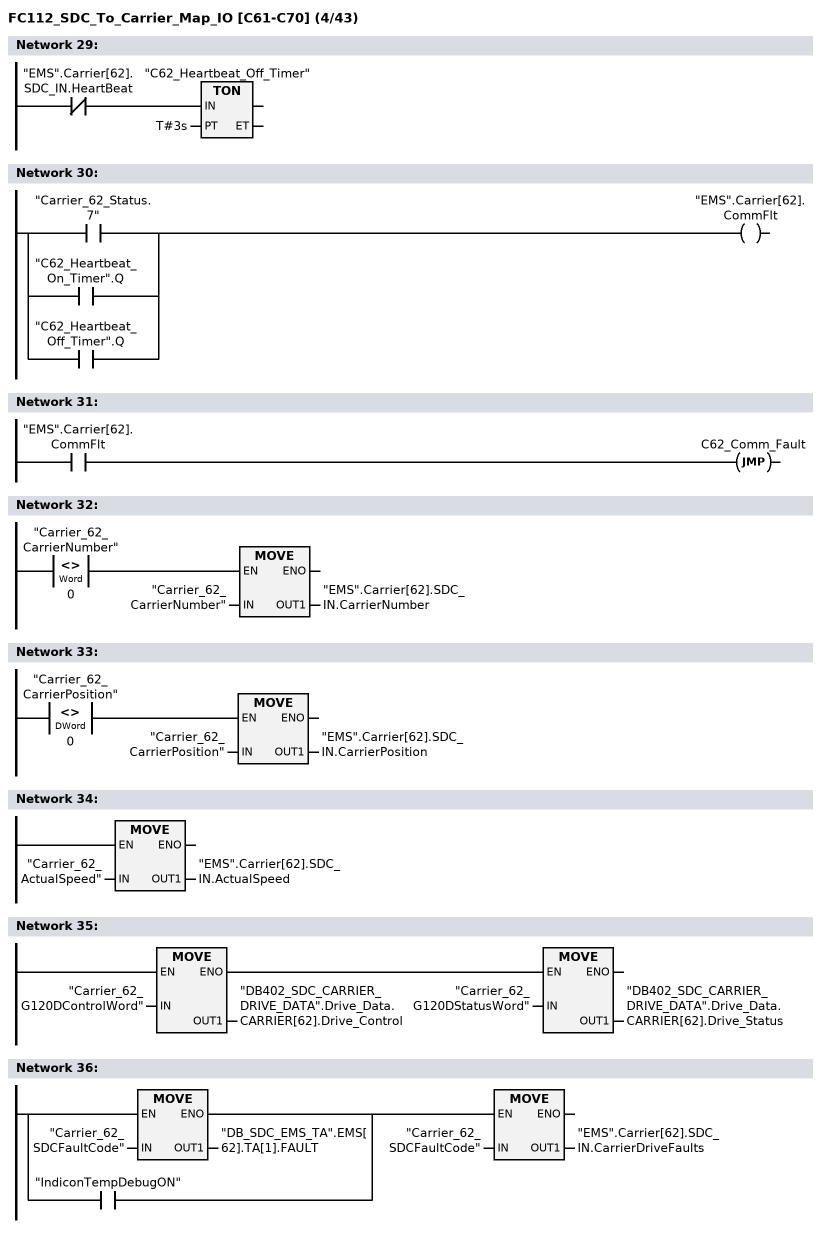
   "C62_Heartbeat_Off_Timer".TON(IN := NOT "EMS".Carrier[62].SDC_IN.HeartBeat, PT := T#3s);
END_REGION

REGION Network 30
   RUNG wire#powerrail
      Contact( "Carrier_62_Status.7" )
      wire#w1
      Coil( "EMS".Carrier[62].CommFlt )
   END_RUNG
   RUNG wire#powerrail
      Contact( "C62_Heartbeat_On_Timer".Q )
   END_RUNG wire#w1
   RUNG wire#powerrail
      Contact( "C62_Heartbeat_Off_Timer".Q )
   END_RUNG wire#w1
   // the same network as SCL:
   "EMS".Carrier[62].CommFlt := "Carrier_62_Status.7" OR "C62_Heartbeat_On_Timer".Q OR "C62_Heartbeat_Off_Timer".Q;
END_REGION

REGION Network 31
   RUNG wire#powerrail
      Contact( "EMS".Carrier[62].CommFlt )
      JumpCoil( C62_Comm_Fault )
   END_RUNG
   // the same network as SCL:
   IF "EMS".Carrier[62].CommFlt THEN GOTO C62_Comm_Fault; END_IF;
END_REGION

REGION Network 32
   RUNG wire#powerrail
      { S7_Templates := "SrcType := Word" } NE_Contact(in1 := "Carrier_62_CarrierNumber", in2 := 0)
      Move(in := "Carrier_62_CarrierNumber", out1 => "EMS".Carrier[62].SDC_IN.CarrierNumber)
   END_RUNG
   // the same network as SCL:
   IF "Carrier_62_CarrierNumber" <> 0 THEN
       "EMS".Carrier[62].SDC_IN.CarrierNumber := "Carrier_62_CarrierNumber";
   END_IF;
END_REGION

REGION Network 33
   RUNG wire#powerrail
      { S7_Templates := "SrcType := DWord" } NE_Contact(in1 := "Carrier_62_CarrierPosition", in2 := 0)
      Move(in := "Carrier_62_CarrierPosition", out1 => "EMS".Carrier[62].SDC_IN.CarrierPosition)
   END_RUNG
   // the same network as SCL:
   IF "Carrier_62_CarrierPosition" <> 0 THEN
       "EMS".Carrier[62].SDC_IN.CarrierPosition := "Carrier_62_CarrierPosition";
   END_IF;
END_REGION

REGION Network 34
   RUNG wire#powerrail
      Move(in := "Carrier_62_ActualSpeed", out1 => "EMS".Carrier[62].SDC_IN.ActualSpeed)
   END_RUNG
   // the same network as SCL:
   "EMS".Carrier[62].SDC_IN.ActualSpeed := "Carrier_62_ActualSpeed";
END_REGION

REGION Network 35
   RUNG wire#powerrail
      Move(in := "Carrier_62_G120DControlWord", out1 => "DB402_SDC_CARRIER_DRIVE_DATA".Drive_Data.CARRIER[62].Drive_Control)
      Move(in := "Carrier_62_G120DStatusWord", out1 => "DB402_SDC_CARRIER_DRIVE_DATA".Drive_Data.CARRIER[62].Drive_Status)
   END_RUNG
   // the same network as SCL:
   "DB402_SDC_CARRIER_DRIVE_DATA".Drive_Data.CARRIER[62].Drive_Control := "Carrier_62_G120DControlWord";
   "DB402_SDC_CARRIER_DRIVE_DATA".Drive_Data.CARRIER[62].Drive_Status := "Carrier_62_G120DStatusWord";
END_REGION

REGION Network 36
   RUNG wire#powerrail
      Move(in := "Carrier_62_SDCFaultCode", out1 => "DB_SDC_EMS_TA".EMS[62].TA[1].FAULT)
      wire#w1
      Move(in := "Carrier_62_SDCFaultCode", out1 => "EMS".Carrier[62].SDC_IN.CarrierDriveFaults)
   END_RUNG
   RUNG wire#powerrail
      Contact( "IndiconTempDebugON" )
   END_RUNG wire#w1
   // the same network as SCL:
   "DB_SDC_EMS_TA".EMS[62].TA[1].FAULT := "Carrier_62_SDCFaultCode";
   IF TRUE OR "IndiconTempDebugON" THEN
       "EMS".Carrier[62].SDC_IN.CarrierDriveFaults := "Carrier_62_SDCFaultCode";
   END_IF;
END_REGION

REGION Network 37
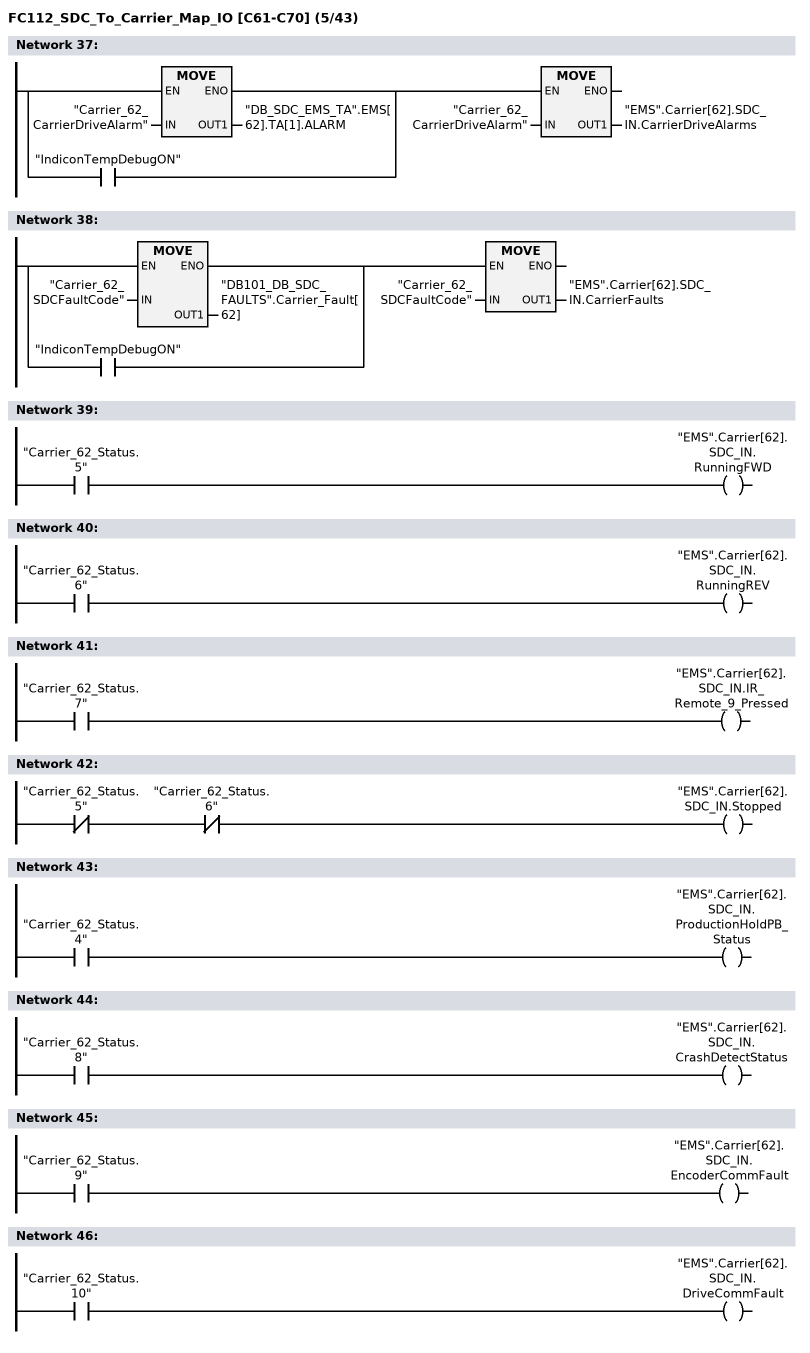
   RUNG wire#powerrail
      Move(in := "Carrier_62_CarrierDriveAlarm", out1 => "DB_SDC_EMS_TA".EMS[62].TA[1].ALARM)
      wire#w1
      Move(in := "Carrier_62_CarrierDriveAlarm", out1 => "EMS".Carrier[62].SDC_IN.CarrierDriveAlarms)
   END_RUNG
   RUNG wire#powerrail
      Contact( "IndiconTempDebugON" )
   END_RUNG wire#w1
   // the same network as SCL:
   "DB_SDC_EMS_TA".EMS[62].TA[1].ALARM := "Carrier_62_CarrierDriveAlarm";
   IF TRUE OR "IndiconTempDebugON" THEN
       "EMS".Carrier[62].SDC_IN.CarrierDriveAlarms := "Carrier_62_CarrierDriveAlarm";
   END_IF;
END_REGION

REGION Network 38
   RUNG wire#powerrail
      Move(in := "Carrier_62_SDCFaultCode", out1 => "DB101_DB_SDC_FAULTS".Carrier_Fault[62])
      wire#w1
      Move(in := "Carrier_62_SDCFaultCode", out1 => "EMS".Carrier[62].SDC_IN.CarrierFaults)
   END_RUNG
   RUNG wire#powerrail
      Contact( "IndiconTempDebugON" )
   END_RUNG wire#w1
   // the same network as SCL:
   "DB101_DB_SDC_FAULTS".Carrier_Fault[62] := "Carrier_62_SDCFaultCode";
   IF TRUE OR "IndiconTempDebugON" THEN
       "EMS".Carrier[62].SDC_IN.CarrierFaults := "Carrier_62_SDCFaultCode";
   END_IF;
END_REGION

REGION Network 39
   RUNG wire#powerrail
      Contact( "Carrier_62_Status.5" )
      Coil( "EMS".Carrier[62].SDC_IN.RunningFWD )
   END_RUNG
   // the same network as SCL:
   "EMS".Carrier[62].SDC_IN.RunningFWD := "Carrier_62_Status.5";
END_REGION

REGION Network 40
   RUNG wire#powerrail
      Contact( "Carrier_62_Status.6" )
      Coil( "EMS".Carrier[62].SDC_IN.RunningREV )
   END_RUNG
   // the same network as SCL:
   "EMS".Carrier[62].SDC_IN.RunningREV := "Carrier_62_Status.6";
END_REGION

REGION Network 41
   RUNG wire#powerrail
      Contact( "Carrier_62_Status.7" )
      Coil( "EMS".Carrier[62].SDC_IN.IR_Remote_9_Pressed )
   END_RUNG
   // the same network as SCL:
   "EMS".Carrier[62].SDC_IN.IR_Remote_9_Pressed := "Carrier_62_Status.7";
END_REGION

REGION Network 42
   RUNG wire#powerrail
      I_Contact( "Carrier_62_Status.5" )
      I_Contact( "Carrier_62_Status.6" )
      Coil( "EMS".Carrier[62].SDC_IN.Stopped )
   END_RUNG
   // the same network as SCL:
   "EMS".Carrier[62].SDC_IN.Stopped := NOT "Carrier_62_Status.5" AND NOT "Carrier_62_Status.6";
END_REGION

REGION Network 43
   RUNG wire#powerrail
      Contact( "Carrier_62_Status.4" )
      Coil( "EMS".Carrier[62].SDC_IN.ProductionHoldPB_Status )
   END_RUNG
   // the same network as SCL:
   "EMS".Carrier[62].SDC_IN.ProductionHoldPB_Status := "Carrier_62_Status.4";
END_REGION

REGION Network 44
   RUNG wire#powerrail
      Contact( "Carrier_62_Status.8" )
      Coil( "EMS".Carrier[62].SDC_IN.CrashDetectStatus )
   END_RUNG
   // the same network as SCL:
   "EMS".Carrier[62].SDC_IN.CrashDetectStatus := "Carrier_62_Status.8";
END_REGION

REGION Network 45
   RUNG wire#powerrail
      Contact( "Carrier_62_Status.9" )
      Coil( "EMS".Carrier[62].SDC_IN.EncoderCommFault )
   END_RUNG
   // the same network as SCL:
   "EMS".Carrier[62].SDC_IN.EncoderCommFault := "Carrier_62_Status.9";
END_REGION

REGION Network 46
   RUNG wire#powerrail
      Contact( "Carrier_62_Status.10" )
      Coil( "EMS".Carrier[62].SDC_IN.DriveCommFault )
   END_RUNG
   // the same network as SCL:
   "EMS".Carrier[62].SDC_IN.DriveCommFault := "Carrier_62_Status.10";
END_REGION

REGION Network 47
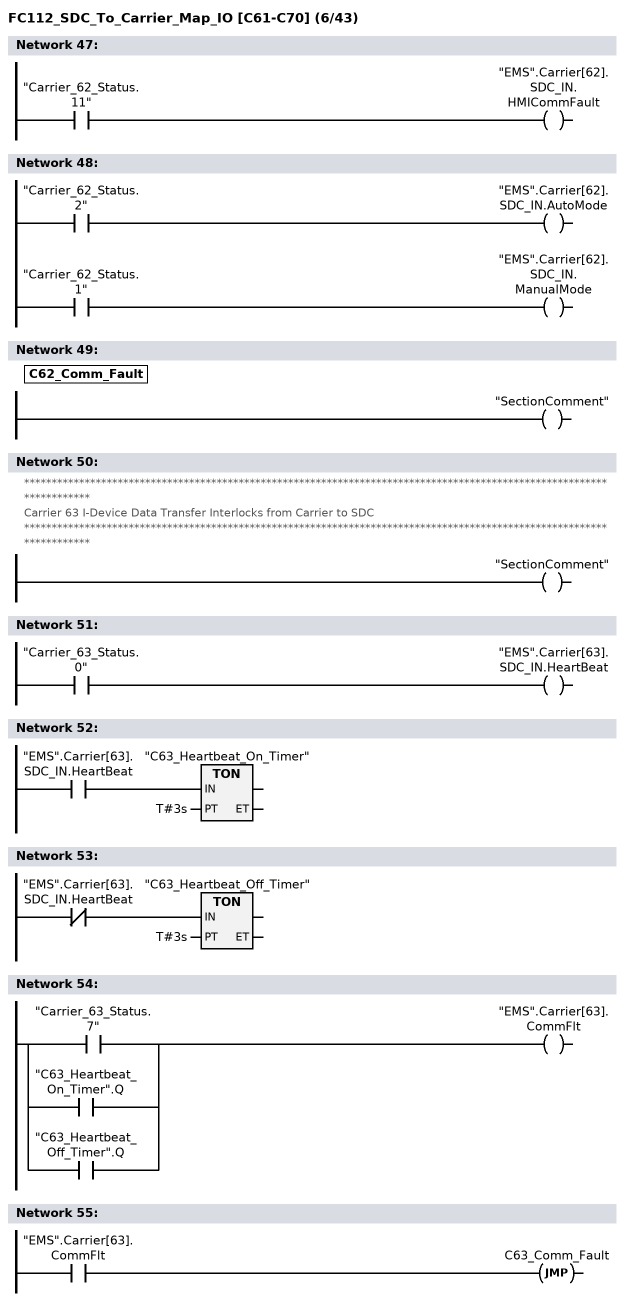
   RUNG wire#powerrail
      Contact( "Carrier_62_Status.11" )
      Coil( "EMS".Carrier[62].SDC_IN.HMICommFault )
   END_RUNG
   // the same network as SCL:
   "EMS".Carrier[62].SDC_IN.HMICommFault := "Carrier_62_Status.11";
END_REGION

REGION Network 48
   RUNG wire#powerrail
      Contact( "Carrier_62_Status.2" )
      Coil( "EMS".Carrier[62].SDC_IN.AutoMode )
   END_RUNG
   RUNG wire#powerrail
      Contact( "Carrier_62_Status.1" )
      Coil( "EMS".Carrier[62].SDC_IN.ManualMode )
   END_RUNG
   // the same network as SCL:
   "EMS".Carrier[62].SDC_IN.AutoMode := "Carrier_62_Status.2";
   "EMS".Carrier[62].SDC_IN.ManualMode := "Carrier_62_Status.1";
END_REGION

REGION Network 49
   Label( C62_Comm_Fault )
   RUNG wire#powerrail
      Coil( "SectionComment" )
   END_RUNG
   // the same network as SCL:
   C62_Comm_Fault:
   "SectionComment" := TRUE;
END_REGION

REGION Network 50
   // **********************************************************************************************************************
   // 
   // Carrier 63 I-Device Data Transfer Interlocks from Carrier to SDC
   // 
   // **********************************************************************************************************************
   RUNG wire#powerrail
      Coil( "SectionComment" )
   END_RUNG
   // the same network as SCL:
   "SectionComment" := TRUE;
END_REGION

REGION Network 51
   RUNG wire#powerrail
      Contact( "Carrier_63_Status.0" )
      Coil( "EMS".Carrier[63].SDC_IN.HeartBeat )
   END_RUNG
   // the same network as SCL:
   "EMS".Carrier[63].SDC_IN.HeartBeat := "Carrier_63_Status.0";
END_REGION

REGION Network 52
   "C63_Heartbeat_On_Timer".TON(IN := "EMS".Carrier[63].SDC_IN.HeartBeat, PT := T#3s);
END_REGION

REGION Network 53
   "C63_Heartbeat_Off_Timer".TON(IN := NOT "EMS".Carrier[63].SDC_IN.HeartBeat, PT := T#3s);
END_REGION

REGION Network 54
   RUNG wire#powerrail
      Contact( "Carrier_63_Status.7" )
      wire#w1
      Coil( "EMS".Carrier[63].CommFlt )
   END_RUNG
   RUNG wire#powerrail
      Contact( "C63_Heartbeat_On_Timer".Q )
   END_RUNG wire#w1
   RUNG wire#powerrail
      Contact( "C63_Heartbeat_Off_Timer".Q )
   END_RUNG wire#w1
   // the same network as SCL:
   "EMS".Carrier[63].CommFlt := "Carrier_63_Status.7" OR "C63_Heartbeat_On_Timer".Q OR "C63_Heartbeat_Off_Timer".Q;
END_REGION

REGION Network 55
   RUNG wire#powerrail
      Contact( "EMS".Carrier[63].CommFlt )
      JumpCoil( C63_Comm_Fault )
   END_RUNG
   // the same network as SCL:
   IF "EMS".Carrier[63].CommFlt THEN GOTO C63_Comm_Fault; END_IF;
END_REGION

REGION Network 56
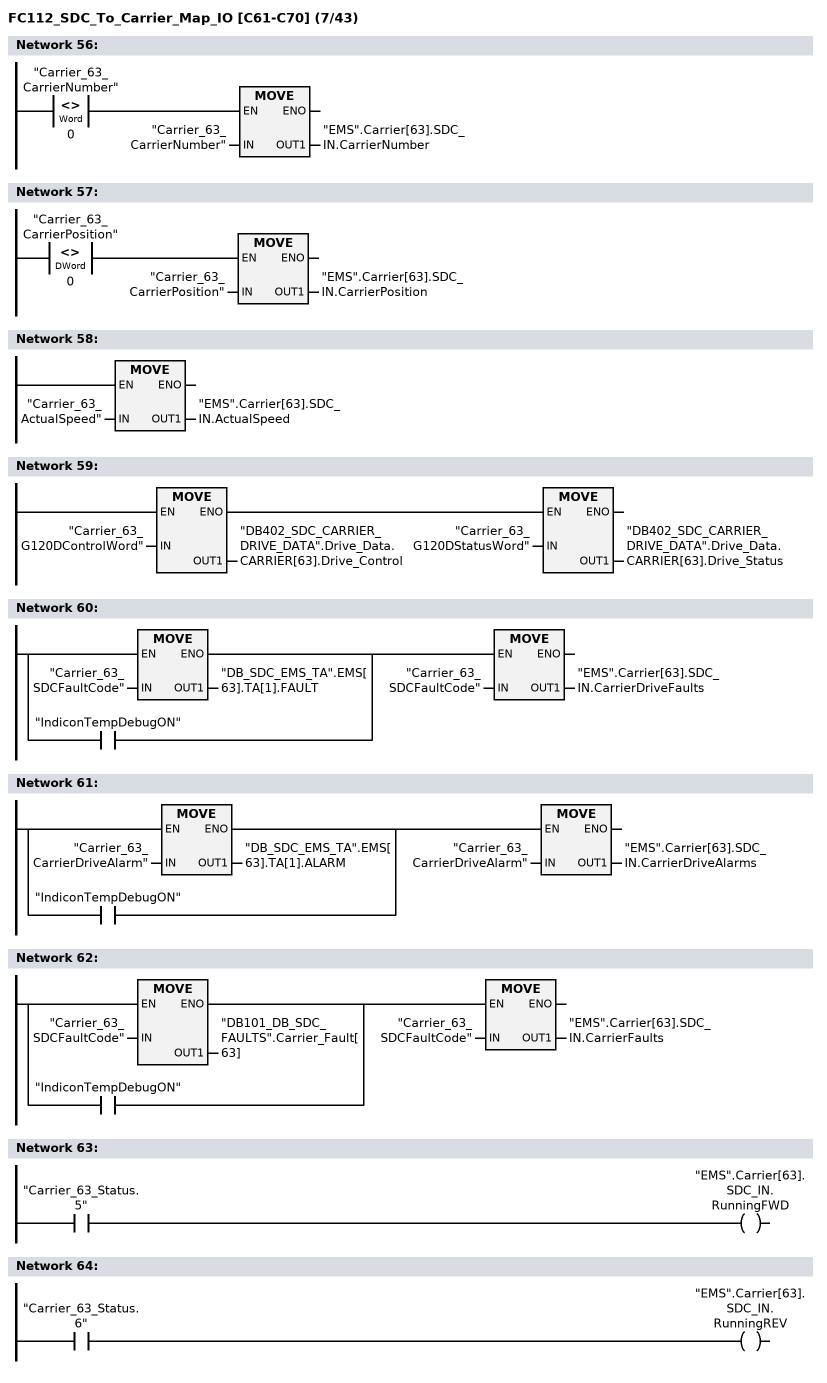
   RUNG wire#powerrail
      { S7_Templates := "SrcType := Word" } NE_Contact(in1 := "Carrier_63_CarrierNumber", in2 := 0)
      Move(in := "Carrier_63_CarrierNumber", out1 => "EMS".Carrier[63].SDC_IN.CarrierNumber)
   END_RUNG
   // the same network as SCL:
   IF "Carrier_63_CarrierNumber" <> 0 THEN
       "EMS".Carrier[63].SDC_IN.CarrierNumber := "Carrier_63_CarrierNumber";
   END_IF;
END_REGION

REGION Network 57
   RUNG wire#powerrail
      { S7_Templates := "SrcType := DWord" } NE_Contact(in1 := "Carrier_63_CarrierPosition", in2 := 0)
      Move(in := "Carrier_63_CarrierPosition", out1 => "EMS".Carrier[63].SDC_IN.CarrierPosition)
   END_RUNG
   // the same network as SCL:
   IF "Carrier_63_CarrierPosition" <> 0 THEN
       "EMS".Carrier[63].SDC_IN.CarrierPosition := "Carrier_63_CarrierPosition";
   END_IF;
END_REGION

REGION Network 58
   RUNG wire#powerrail
      Move(in := "Carrier_63_ActualSpeed", out1 => "EMS".Carrier[63].SDC_IN.ActualSpeed)
   END_RUNG
   // the same network as SCL:
   "EMS".Carrier[63].SDC_IN.ActualSpeed := "Carrier_63_ActualSpeed";
END_REGION

REGION Network 59
   RUNG wire#powerrail
      Move(in := "Carrier_63_G120DControlWord", out1 => "DB402_SDC_CARRIER_DRIVE_DATA".Drive_Data.CARRIER[63].Drive_Control)
      Move(in := "Carrier_63_G120DStatusWord", out1 => "DB402_SDC_CARRIER_DRIVE_DATA".Drive_Data.CARRIER[63].Drive_Status)
   END_RUNG
   // the same network as SCL:
   "DB402_SDC_CARRIER_DRIVE_DATA".Drive_Data.CARRIER[63].Drive_Control := "Carrier_63_G120DControlWord";
   "DB402_SDC_CARRIER_DRIVE_DATA".Drive_Data.CARRIER[63].Drive_Status := "Carrier_63_G120DStatusWord";
END_REGION

REGION Network 60
   RUNG wire#powerrail
      Move(in := "Carrier_63_SDCFaultCode", out1 => "DB_SDC_EMS_TA".EMS[63].TA[1].FAULT)
      wire#w1
      Move(in := "Carrier_63_SDCFaultCode", out1 => "EMS".Carrier[63].SDC_IN.CarrierDriveFaults)
   END_RUNG
   RUNG wire#powerrail
      Contact( "IndiconTempDebugON" )
   END_RUNG wire#w1
   // the same network as SCL:
   "DB_SDC_EMS_TA".EMS[63].TA[1].FAULT := "Carrier_63_SDCFaultCode";
   IF TRUE OR "IndiconTempDebugON" THEN
       "EMS".Carrier[63].SDC_IN.CarrierDriveFaults := "Carrier_63_SDCFaultCode";
   END_IF;
END_REGION

REGION Network 61
   RUNG wire#powerrail
      Move(in := "Carrier_63_CarrierDriveAlarm", out1 => "DB_SDC_EMS_TA".EMS[63].TA[1].ALARM)
      wire#w1
      Move(in := "Carrier_63_CarrierDriveAlarm", out1 => "EMS".Carrier[63].SDC_IN.CarrierDriveAlarms)
   END_RUNG
   RUNG wire#powerrail
      Contact( "IndiconTempDebugON" )
   END_RUNG wire#w1
   // the same network as SCL:
   "DB_SDC_EMS_TA".EMS[63].TA[1].ALARM := "Carrier_63_CarrierDriveAlarm";
   IF TRUE OR "IndiconTempDebugON" THEN
       "EMS".Carrier[63].SDC_IN.CarrierDriveAlarms := "Carrier_63_CarrierDriveAlarm";
   END_IF;
END_REGION

REGION Network 62
   RUNG wire#powerrail
      Move(in := "Carrier_63_SDCFaultCode", out1 => "DB101_DB_SDC_FAULTS".Carrier_Fault[63])
      wire#w1
      Move(in := "Carrier_63_SDCFaultCode", out1 => "EMS".Carrier[63].SDC_IN.CarrierFaults)
   END_RUNG
   RUNG wire#powerrail
      Contact( "IndiconTempDebugON" )
   END_RUNG wire#w1
   // the same network as SCL:
   "DB101_DB_SDC_FAULTS".Carrier_Fault[63] := "Carrier_63_SDCFaultCode";
   IF TRUE OR "IndiconTempDebugON" THEN
       "EMS".Carrier[63].SDC_IN.CarrierFaults := "Carrier_63_SDCFaultCode";
   END_IF;
END_REGION

REGION Network 63
   RUNG wire#powerrail
      Contact( "Carrier_63_Status.5" )
      Coil( "EMS".Carrier[63].SDC_IN.RunningFWD )
   END_RUNG
   // the same network as SCL:
   "EMS".Carrier[63].SDC_IN.RunningFWD := "Carrier_63_Status.5";
END_REGION

REGION Network 64
   RUNG wire#powerrail
      Contact( "Carrier_63_Status.6" )
      Coil( "EMS".Carrier[63].SDC_IN.RunningREV )
   END_RUNG
   // the same network as SCL:
   "EMS".Carrier[63].SDC_IN.RunningREV := "Carrier_63_Status.6";
END_REGION

REGION Network 65
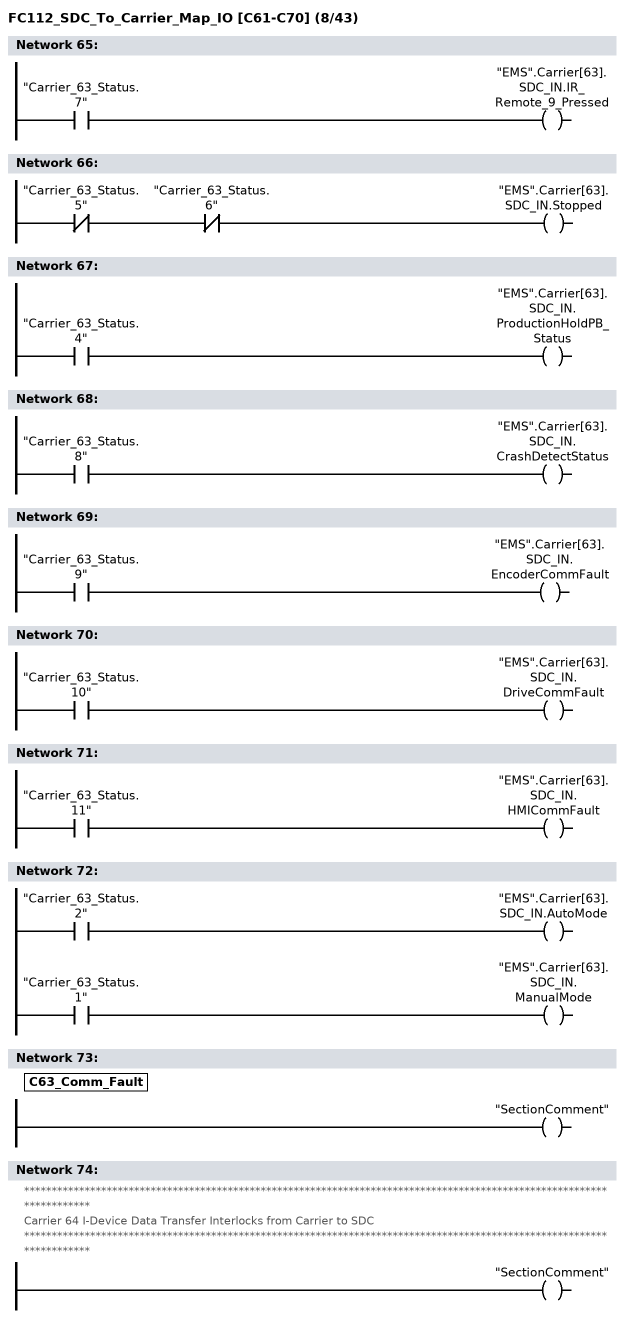
   RUNG wire#powerrail
      Contact( "Carrier_63_Status.7" )
      Coil( "EMS".Carrier[63].SDC_IN.IR_Remote_9_Pressed )
   END_RUNG
   // the same network as SCL:
   "EMS".Carrier[63].SDC_IN.IR_Remote_9_Pressed := "Carrier_63_Status.7";
END_REGION

REGION Network 66
   RUNG wire#powerrail
      I_Contact( "Carrier_63_Status.5" )
      I_Contact( "Carrier_63_Status.6" )
      Coil( "EMS".Carrier[63].SDC_IN.Stopped )
   END_RUNG
   // the same network as SCL:
   "EMS".Carrier[63].SDC_IN.Stopped := NOT "Carrier_63_Status.5" AND NOT "Carrier_63_Status.6";
END_REGION

REGION Network 67
   RUNG wire#powerrail
      Contact( "Carrier_63_Status.4" )
      Coil( "EMS".Carrier[63].SDC_IN.ProductionHoldPB_Status )
   END_RUNG
   // the same network as SCL:
   "EMS".Carrier[63].SDC_IN.ProductionHoldPB_Status := "Carrier_63_Status.4";
END_REGION

REGION Network 68
   RUNG wire#powerrail
      Contact( "Carrier_63_Status.8" )
      Coil( "EMS".Carrier[63].SDC_IN.CrashDetectStatus )
   END_RUNG
   // the same network as SCL:
   "EMS".Carrier[63].SDC_IN.CrashDetectStatus := "Carrier_63_Status.8";
END_REGION

REGION Network 69
   RUNG wire#powerrail
      Contact( "Carrier_63_Status.9" )
      Coil( "EMS".Carrier[63].SDC_IN.EncoderCommFault )
   END_RUNG
   // the same network as SCL:
   "EMS".Carrier[63].SDC_IN.EncoderCommFault := "Carrier_63_Status.9";
END_REGION

REGION Network 70
   RUNG wire#powerrail
      Contact( "Carrier_63_Status.10" )
      Coil( "EMS".Carrier[63].SDC_IN.DriveCommFault )
   END_RUNG
   // the same network as SCL:
   "EMS".Carrier[63].SDC_IN.DriveCommFault := "Carrier_63_Status.10";
END_REGION

REGION Network 71
   RUNG wire#powerrail
      Contact( "Carrier_63_Status.11" )
      Coil( "EMS".Carrier[63].SDC_IN.HMICommFault )
   END_RUNG
   // the same network as SCL:
   "EMS".Carrier[63].SDC_IN.HMICommFault := "Carrier_63_Status.11";
END_REGION

REGION Network 72
   RUNG wire#powerrail
      Contact( "Carrier_63_Status.2" )
      Coil( "EMS".Carrier[63].SDC_IN.AutoMode )
   END_RUNG
   RUNG wire#powerrail
      Contact( "Carrier_63_Status.1" )
      Coil( "EMS".Carrier[63].SDC_IN.ManualMode )
   END_RUNG
   // the same network as SCL:
   "EMS".Carrier[63].SDC_IN.AutoMode := "Carrier_63_Status.2";
   "EMS".Carrier[63].SDC_IN.ManualMode := "Carrier_63_Status.1";
END_REGION

REGION Network 73
   Label( C63_Comm_Fault )
   RUNG wire#powerrail
      Coil( "SectionComment" )
   END_RUNG
   // the same network as SCL:
   C63_Comm_Fault:
   "SectionComment" := TRUE;
END_REGION

REGION Network 74
   // **********************************************************************************************************************
   // 
   // Carrier 64 I-Device Data Transfer Interlocks from Carrier to SDC
   // 
   // **********************************************************************************************************************
   RUNG wire#powerrail
      Coil( "SectionComment" )
   END_RUNG
   // the same network as SCL:
   "SectionComment" := TRUE;
END_REGION

REGION Network 75
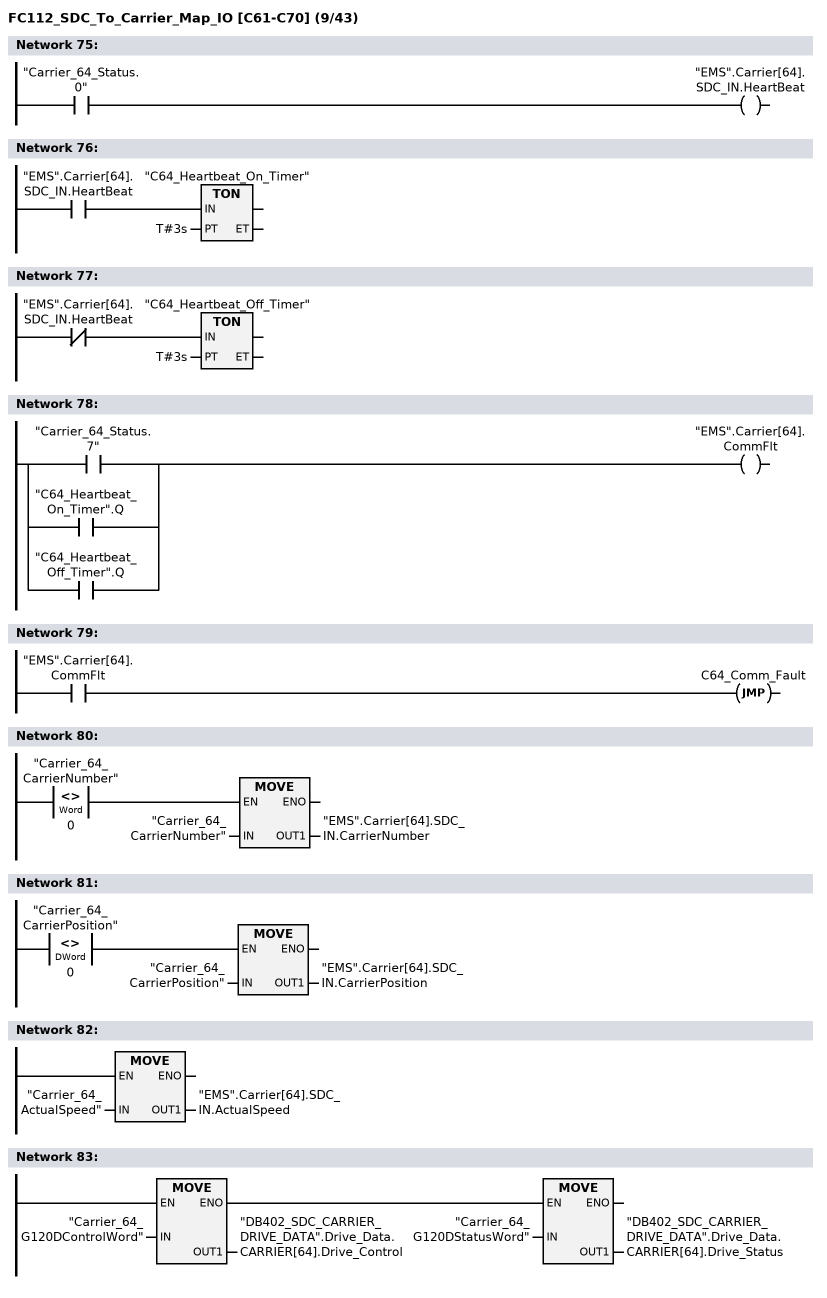
   RUNG wire#powerrail
      Contact( "Carrier_64_Status.0" )
      Coil( "EMS".Carrier[64].SDC_IN.HeartBeat )
   END_RUNG
   // the same network as SCL:
   "EMS".Carrier[64].SDC_IN.HeartBeat := "Carrier_64_Status.0";
END_REGION

REGION Network 76
   "C64_Heartbeat_On_Timer".TON(IN := "EMS".Carrier[64].SDC_IN.HeartBeat, PT := T#3s);
END_REGION

REGION Network 77
   "C64_Heartbeat_Off_Timer".TON(IN := NOT "EMS".Carrier[64].SDC_IN.HeartBeat, PT := T#3s);
END_REGION

REGION Network 78
   RUNG wire#powerrail
      Contact( "Carrier_64_Status.7" )
      wire#w1
      Coil( "EMS".Carrier[64].CommFlt )
   END_RUNG
   RUNG wire#powerrail
      Contact( "C64_Heartbeat_On_Timer".Q )
   END_RUNG wire#w1
   RUNG wire#powerrail
      Contact( "C64_Heartbeat_Off_Timer".Q )
   END_RUNG wire#w1
   // the same network as SCL:
   "EMS".Carrier[64].CommFlt := "Carrier_64_Status.7" OR "C64_Heartbeat_On_Timer".Q OR "C64_Heartbeat_Off_Timer".Q;
END_REGION

REGION Network 79
   RUNG wire#powerrail
      Contact( "EMS".Carrier[64].CommFlt )
      JumpCoil( C64_Comm_Fault )
   END_RUNG
   // the same network as SCL:
   IF "EMS".Carrier[64].CommFlt THEN GOTO C64_Comm_Fault; END_IF;
END_REGION

REGION Network 80
   RUNG wire#powerrail
      { S7_Templates := "SrcType := Word" } NE_Contact(in1 := "Carrier_64_CarrierNumber", in2 := 0)
      Move(in := "Carrier_64_CarrierNumber", out1 => "EMS".Carrier[64].SDC_IN.CarrierNumber)
   END_RUNG
   // the same network as SCL:
   IF "Carrier_64_CarrierNumber" <> 0 THEN
       "EMS".Carrier[64].SDC_IN.CarrierNumber := "Carrier_64_CarrierNumber";
   END_IF;
END_REGION

REGION Network 81
   RUNG wire#powerrail
      { S7_Templates := "SrcType := DWord" } NE_Contact(in1 := "Carrier_64_CarrierPosition", in2 := 0)
      Move(in := "Carrier_64_CarrierPosition", out1 => "EMS".Carrier[64].SDC_IN.CarrierPosition)
   END_RUNG
   // the same network as SCL:
   IF "Carrier_64_CarrierPosition" <> 0 THEN
       "EMS".Carrier[64].SDC_IN.CarrierPosition := "Carrier_64_CarrierPosition";
   END_IF;
END_REGION

REGION Network 82
   RUNG wire#powerrail
      Move(in := "Carrier_64_ActualSpeed", out1 => "EMS".Carrier[64].SDC_IN.ActualSpeed)
   END_RUNG
   // the same network as SCL:
   "EMS".Carrier[64].SDC_IN.ActualSpeed := "Carrier_64_ActualSpeed";
END_REGION

REGION Network 83
   RUNG wire#powerrail
      Move(in := "Carrier_64_G120DControlWord", out1 => "DB402_SDC_CARRIER_DRIVE_DATA".Drive_Data.CARRIER[64].Drive_Control)
      Move(in := "Carrier_64_G120DStatusWord", out1 => "DB402_SDC_CARRIER_DRIVE_DATA".Drive_Data.CARRIER[64].Drive_Status)
   END_RUNG
   // the same network as SCL:
   "DB402_SDC_CARRIER_DRIVE_DATA".Drive_Data.CARRIER[64].Drive_Control := "Carrier_64_G120DControlWord";
   "DB402_SDC_CARRIER_DRIVE_DATA".Drive_Data.CARRIER[64].Drive_Status := "Carrier_64_G120DStatusWord";
END_REGION

REGION Network 84
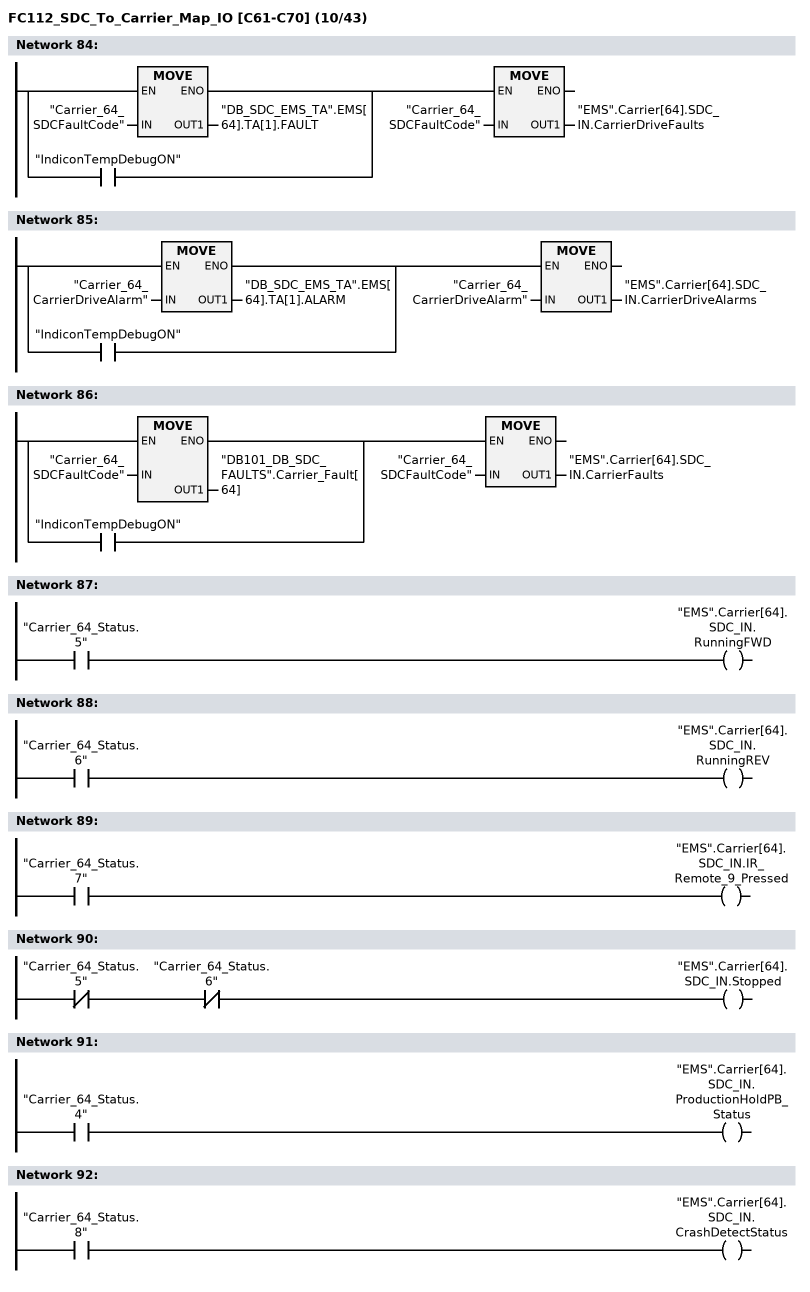
   RUNG wire#powerrail
      Move(in := "Carrier_64_SDCFaultCode", out1 => "DB_SDC_EMS_TA".EMS[64].TA[1].FAULT)
      wire#w1
      Move(in := "Carrier_64_SDCFaultCode", out1 => "EMS".Carrier[64].SDC_IN.CarrierDriveFaults)
   END_RUNG
   RUNG wire#powerrail
      Contact( "IndiconTempDebugON" )
   END_RUNG wire#w1
   // the same network as SCL:
   "DB_SDC_EMS_TA".EMS[64].TA[1].FAULT := "Carrier_64_SDCFaultCode";
   IF TRUE OR "IndiconTempDebugON" THEN
       "EMS".Carrier[64].SDC_IN.CarrierDriveFaults := "Carrier_64_SDCFaultCode";
   END_IF;
END_REGION

REGION Network 85
   RUNG wire#powerrail
      Move(in := "Carrier_64_CarrierDriveAlarm", out1 => "DB_SDC_EMS_TA".EMS[64].TA[1].ALARM)
      wire#w1
      Move(in := "Carrier_64_CarrierDriveAlarm", out1 => "EMS".Carrier[64].SDC_IN.CarrierDriveAlarms)
   END_RUNG
   RUNG wire#powerrail
      Contact( "IndiconTempDebugON" )
   END_RUNG wire#w1
   // the same network as SCL:
   "DB_SDC_EMS_TA".EMS[64].TA[1].ALARM := "Carrier_64_CarrierDriveAlarm";
   IF TRUE OR "IndiconTempDebugON" THEN
       "EMS".Carrier[64].SDC_IN.CarrierDriveAlarms := "Carrier_64_CarrierDriveAlarm";
   END_IF;
END_REGION

REGION Network 86
   RUNG wire#powerrail
      Move(in := "Carrier_64_SDCFaultCode", out1 => "DB101_DB_SDC_FAULTS".Carrier_Fault[64])
      wire#w1
      Move(in := "Carrier_64_SDCFaultCode", out1 => "EMS".Carrier[64].SDC_IN.CarrierFaults)
   END_RUNG
   RUNG wire#powerrail
      Contact( "IndiconTempDebugON" )
   END_RUNG wire#w1
   // the same network as SCL:
   "DB101_DB_SDC_FAULTS".Carrier_Fault[64] := "Carrier_64_SDCFaultCode";
   IF TRUE OR "IndiconTempDebugON" THEN
       "EMS".Carrier[64].SDC_IN.CarrierFaults := "Carrier_64_SDCFaultCode";
   END_IF;
END_REGION

REGION Network 87
   RUNG wire#powerrail
      Contact( "Carrier_64_Status.5" )
      Coil( "EMS".Carrier[64].SDC_IN.RunningFWD )
   END_RUNG
   // the same network as SCL:
   "EMS".Carrier[64].SDC_IN.RunningFWD := "Carrier_64_Status.5";
END_REGION

REGION Network 88
   RUNG wire#powerrail
      Contact( "Carrier_64_Status.6" )
      Coil( "EMS".Carrier[64].SDC_IN.RunningREV )
   END_RUNG
   // the same network as SCL:
   "EMS".Carrier[64].SDC_IN.RunningREV := "Carrier_64_Status.6";
END_REGION

REGION Network 89
   RUNG wire#powerrail
      Contact( "Carrier_64_Status.7" )
      Coil( "EMS".Carrier[64].SDC_IN.IR_Remote_9_Pressed )
   END_RUNG
   // the same network as SCL:
   "EMS".Carrier[64].SDC_IN.IR_Remote_9_Pressed := "Carrier_64_Status.7";
END_REGION

REGION Network 90
   RUNG wire#powerrail
      I_Contact( "Carrier_64_Status.5" )
      I_Contact( "Carrier_64_Status.6" )
      Coil( "EMS".Carrier[64].SDC_IN.Stopped )
   END_RUNG
   // the same network as SCL:
   "EMS".Carrier[64].SDC_IN.Stopped := NOT "Carrier_64_Status.5" AND NOT "Carrier_64_Status.6";
END_REGION

REGION Network 91
   RUNG wire#powerrail
      Contact( "Carrier_64_Status.4" )
      Coil( "EMS".Carrier[64].SDC_IN.ProductionHoldPB_Status )
   END_RUNG
   // the same network as SCL:
   "EMS".Carrier[64].SDC_IN.ProductionHoldPB_Status := "Carrier_64_Status.4";
END_REGION

REGION Network 92
   RUNG wire#powerrail
      Contact( "Carrier_64_Status.8" )
      Coil( "EMS".Carrier[64].SDC_IN.CrashDetectStatus )
   END_RUNG
   // the same network as SCL:
   "EMS".Carrier[64].SDC_IN.CrashDetectStatus := "Carrier_64_Status.8";
END_REGION

REGION Network 93
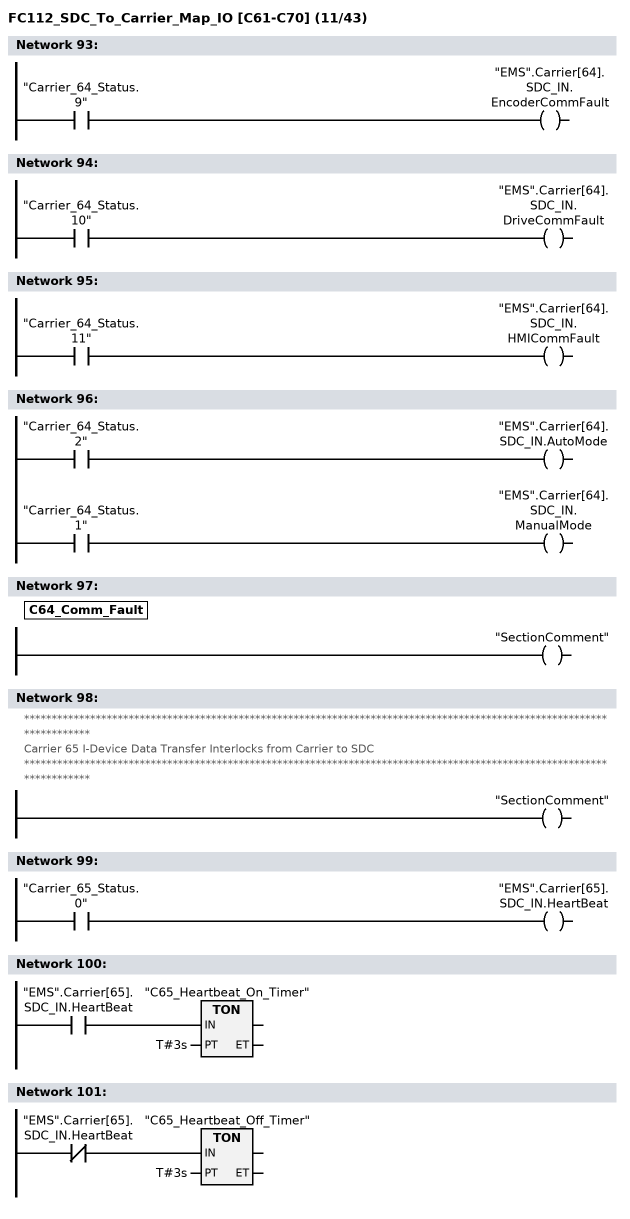
   RUNG wire#powerrail
      Contact( "Carrier_64_Status.9" )
      Coil( "EMS".Carrier[64].SDC_IN.EncoderCommFault )
   END_RUNG
   // the same network as SCL:
   "EMS".Carrier[64].SDC_IN.EncoderCommFault := "Carrier_64_Status.9";
END_REGION

REGION Network 94
   RUNG wire#powerrail
      Contact( "Carrier_64_Status.10" )
      Coil( "EMS".Carrier[64].SDC_IN.DriveCommFault )
   END_RUNG
   // the same network as SCL:
   "EMS".Carrier[64].SDC_IN.DriveCommFault := "Carrier_64_Status.10";
END_REGION

REGION Network 95
   RUNG wire#powerrail
      Contact( "Carrier_64_Status.11" )
      Coil( "EMS".Carrier[64].SDC_IN.HMICommFault )
   END_RUNG
   // the same network as SCL:
   "EMS".Carrier[64].SDC_IN.HMICommFault := "Carrier_64_Status.11";
END_REGION

REGION Network 96
   RUNG wire#powerrail
      Contact( "Carrier_64_Status.2" )
      Coil( "EMS".Carrier[64].SDC_IN.AutoMode )
   END_RUNG
   RUNG wire#powerrail
      Contact( "Carrier_64_Status.1" )
      Coil( "EMS".Carrier[64].SDC_IN.ManualMode )
   END_RUNG
   // the same network as SCL:
   "EMS".Carrier[64].SDC_IN.AutoMode := "Carrier_64_Status.2";
   "EMS".Carrier[64].SDC_IN.ManualMode := "Carrier_64_Status.1";
END_REGION

REGION Network 97
   Label( C64_Comm_Fault )
   RUNG wire#powerrail
      Coil( "SectionComment" )
   END_RUNG
   // the same network as SCL:
   C64_Comm_Fault:
   "SectionComment" := TRUE;
END_REGION

REGION Network 98
   // **********************************************************************************************************************
   // 
   // Carrier 65 I-Device Data Transfer Interlocks from Carrier to SDC
   // 
   // **********************************************************************************************************************
   RUNG wire#powerrail
      Coil( "SectionComment" )
   END_RUNG
   // the same network as SCL:
   "SectionComment" := TRUE;
END_REGION

REGION Network 99
   RUNG wire#powerrail
      Contact( "Carrier_65_Status.0" )
      Coil( "EMS".Carrier[65].SDC_IN.HeartBeat )
   END_RUNG
   // the same network as SCL:
   "EMS".Carrier[65].SDC_IN.HeartBeat := "Carrier_65_Status.0";
END_REGION

REGION Network 100
   "C65_Heartbeat_On_Timer".TON(IN := "EMS".Carrier[65].SDC_IN.HeartBeat, PT := T#3s);
END_REGION

REGION Network 101
   "C65_Heartbeat_Off_Timer".TON(IN := NOT "EMS".Carrier[65].SDC_IN.HeartBeat, PT := T#3s);
END_REGION

REGION Network 102